
               #STATE_FAULT,
               #STATE_PROBLEM:
                   // The device is reachable, but faulty because of an error in a
                   // subordinated system --> check the modules
                   // Store the state of the different module in the diag DB
                   FOR #tempSlotIndex := 0 TO "USERDIAG_SLOTS_PER_DEVICE_UPPER_LIM" DO
                       IF (#ioSystemData.devices[#tempDeviceIndex].slots[#tempSlotIndex].configured = TRUE)
                       THEN
                           IF (#statDeviceProblemModules[#tempSlotIndex + 1] = TRUE)
                           THEN
                               // Problem in module
                               #ioSystemData.devices[#tempDeviceIndex].slots[#tempSlotIndex].faulty := FALSE;
                               #ioSystemData.devices[#tempDeviceIndex].slots[#tempSlotIndex].error := TRUE;
                               #ioSystemData.devices[#tempDeviceIndex].slots[#tempSlotIndex].problem := TRUE;
                               #ioSystemData.devices[#tempDeviceIndex].slots[#tempSlotIndex].state := #STATE_PROBLEM;

                               IF (#statDeviceFaultyModules[#tempSlotIndex + 1] = TRUE)
                               THEN
                                   // Fault in module
                                   #ioSystemData.devices[#tempDeviceIndex].slots[#tempSlotIndex].faulty := TRUE;
                                   #ioSystemData.devices[#tempDeviceIndex].slots[#tempSlotIndex].state := #STATE_FAULT;
                               END_IF;
                           ELSE
                               #ioSystemData.devices[#tempDeviceIndex].slots[#tempSlotIndex].error := FALSE;
                               #ioSystemData.devices[#tempDeviceIndex].slots[#tempSlotIndex].problem := FALSE;
                               #ioSystemData.devices[#tempDeviceIndex].slots[#tempSlotIndex].faulty := FALSE;
                           END_IF;

                           IF (#statDeviceExistingModules[#tempSlotIndex + 1] = TRUE)
                           THEN
                               // Module exists
                               #ioSystemData.devices[#tempDeviceIndex].slots[#tempSlotIndex].exists := TRUE;
                           ELSE
                               // Module does not exist
                               #ioSystemData.devices[#tempDeviceIndex].slots[#tempSlotIndex].exists := FALSE;
                           END_IF;
                       END_IF;
                   END_FOR;
               ELSE
                   // All modules are okay
                   FOR #tempSlotIndex := 0 TO "USERDIAG_SLOTS_PER_DEVICE_UPPER_LIM" DO
                       IF (#ioSystemData.devices[#tempDeviceIndex].slots[#tempSlotIndex].configured = TRUE)
                       THEN
                           #ioSystemData.devices[#tempDeviceIndex].slots[#tempSlotIndex].error := FALSE;
                           #ioSystemData.devices[#tempDeviceIndex].slots[#tempSlotIndex].problem := FALSE;
                           #ioSystemData.devices[#tempDeviceIndex].slots[#tempSlotIndex].faulty := FALSE;
                           #ioSystemData.devices[#tempDeviceIndex].slots[#tempSlotIndex].exists := TRUE;
                       END_IF;
                   END_FOR;
           END_CASE;
       END_IF;

       // Initialize the pointer for the next run
       #tempDeviceIndex := #ioSystemData.devices[#tempDeviceIndex].nextDevice;
   END_WHILE;


   // Write static values to outputs
   #error := #statError;
   #status := #statStatus;
   #statusID := #statStatusID;
END_FUNCTION_BLOCK

// folder: OBs

ORGANIZATION_BLOCK "Main"   // OB1, LAD, ProgramCycle
TITLE = "Main Program Sweep (Cycle)"
{ S7_Optimized_Access := 'TRUE' }
VERSION : 0.1
   VAR_INPUT
      Initial_Call : Bool;   // Initial call of this OB
      Remanence : Bool;   // =True, if remanent data are available
   END_VAR
BEGIN

REGION Network 1
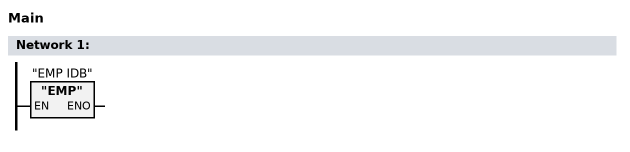
   RUNG wire#powerrail
      "EMP IDB"()
   END_RUNG
   // the same network as SCL:
   "EMP IDB"();   // "EMP"
END_REGION
END_ORGANIZATION_BLOCK

ORGANIZATION_BLOCK "Rack or station failure"   // OB86, LAD, RackStationFailure
{ S7_Optimized_Access := 'TRUE' }
VERSION : 0.1
   VAR_INPUT
      LADDR : Hw_Device;   // Hardware identifier
      Event_Class : Byte;   // Event class
      Fault_ID : Byte;   // Fault identifier
   END_VAR
BEGIN
END_ORGANIZATION_BLOCK

ORGANIZATION_BLOCK "Startup"   // OB100, LAD, Startup
TITLE = "Complete Restart"
{ S7_Optimized_Access := 'TRUE' }
VERSION : 0.1
// //============================================================================
// //SIEMENS AG
// //(c)Copyright 2017 All Rights Reserved
// //-----------------------------------------------------------------------------
// //Library: -
// //Tested with: S7-1516-3 PN/DP FW 2.5
// //Engineering: TIA Portal V15
// //Restrictions: -
// //Requirements: -
// //Functionality: Startup OB for Diagnostics
// //-----------------------------------------------------------------------------
// //Change log table:
// //Version  Date              Expert in charge                               Changes applied
// //01.00.00 25.04.2017 Siemens Industry Online Support First released version
// //============================================================================
   VAR_INPUT
      LostRetentive : Bool;   // True if retentive data are lost
      LostRTC : Bool;   // True if date and time are lost
   END_VAR
   VAR_TEMP
      index : Int;
   END_VAR
BEGIN

REGION Network 1: Set start user diagnostic
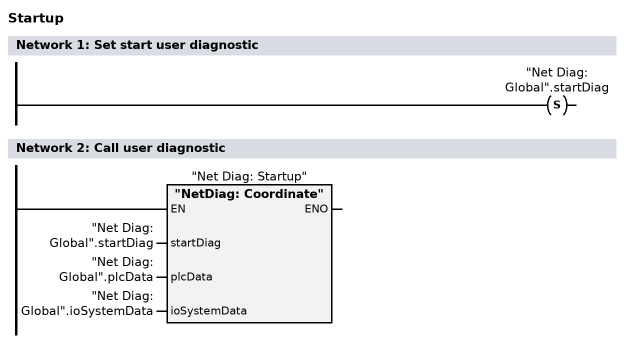
   RUNG wire#powerrail
      S_Coil( "Net Diag: Global".startDiag )
   END_RUNG
   // the same network as SCL:
   "Net Diag: Global".startDiag := TRUE;
END_REGION

REGION Network 2: Call user diagnostic
   RUNG wire#powerrail
      "Net Diag: Startup"(startDiag := "Net Diag: Global".startDiag, plcData := "Net Diag: Global".plcData, ioSystemData := "Net Diag: Global".ioSystemData)
   END_RUNG
   // the same network as SCL:
   "Net Diag: Startup"(startDiag := "Net Diag: Global".startDiag,   // "NetDiag: Coordinate"
                       plcData := "Net Diag: Global".plcData,
                       ioSystemData := "Net Diag: Global".ioSystemData);
END_REGION
END_ORGANIZATION_BLOCK

ORGANIZATION_BLOCK "Programming error"   // OB121, LAD, ProgrammingError
{ S7_Optimized_Access := 'TRUE' }
VERSION : 0.1
   VAR_INPUT
      BlockNr : UInt;   // Number of causing block
      Reaction : USInt;   // 0:ignore, 1:substitute, 2:skip
      Fault_ID : Byte;   // Fault identifier
      BlockType : USInt;   // 16#01:OB, 16#02:FC, 16#03:FB, 16#04:SFC, 16#05:SFB, 16#06:DB: Type of block causing the error
      Area : USInt;   // Area where the error occured
      DBNr : DB_ANY;   // DB number if Area = DB or DI
      Csg_OBNr : OB_Any;   // Number of OB causing the error
      Csg_Prio : USInt;   // Priority of OB causing the error
      Width : USInt;   // 0:bit, 1:byte, 2:word, 3:dword, 4:lword
   END_VAR
BEGIN
END_ORGANIZATION_BLOCK

ORGANIZATION_BLOCK "IO access error"   // OB122, LAD, IOAccessError
{ S7_Optimized_Access := 'TRUE' }
VERSION : 0.1
   VAR_INPUT
      BlockNr : UInt;   // Number of causing block
      Reaction : USInt;   // 0:ignore, 1:substitute, 2:skip
      Fault_ID : Byte;   // 16#42:reading, 16#43:writing
      BlockType : USInt;   // 16#01:OB, 16#02:FC, 16#03:FB, 16#04:SFC, 16#05:SFB, 16#06:DB: Type of block causing the error
      Area : USInt;   // 16#81:I, 16#82:Q: IO area where the IOaccess error occured
      DBNr : DB_ANY;   // Reserved for system
      Csg_OBNr : OB_Any;   // Number of OB causing the error
      Csg_Prio : USInt;   // Priority of OB causing the error
      Width : USInt;   // 0:bit, 1:byte, 2:word, 3:dword, 4:lword
   END_VAR
BEGIN
END_ORGANIZATION_BLOCK

// folder: Unsorted

FUNCTION_BLOCK "Code 128"   // FB2, SCL
{ S7_Optimized_Access := 'TRUE' }
VERSION : 0.1
   VAR_INPUT
      partNumber : String;
   END_VAR
   VAR_OUTPUT
      barcode : String;
   END_VAR
   VAR
      charsIn : Array[0..255] of Byte;
      charsOut : Array[0..255] of Byte;
      cnt : UInt;
      intVals : Array[0..255] of Int;
      sum : Int;
      checkSum : Int;
   END_VAR
   VAR_TEMP
      pn : String;
      i : Int;
   END_VAR
   VAR CONSTANT
      startChar : Char := 'Ì';
      stopChar : Char := 'Î';
   END_VAR
   // intVals[0] := 104;
BEGIN
   #pn := #partNumber;

   FOR #i := 0 TO 255 DO
       #charsIn[#i] := 16#00;
       #charsOut[#i] := 16#00;
       #intVals[#i] := 0;
   END_FOR;

   Strg_TO_Chars(Strg:=#pn,
                 pChars:=0,
                 Cnt=>#cnt,
                 Chars:=#charsIn);


   #sum := 104;
   FOR #i := 0 TO UINT_TO_INT(#cnt - 1) DO
       #intVals[#i] := CHAR_TO_INT(#charsIn[#i]) - 32;
       #intVals[#i] := #intVals[#i] * (#i + 1);
       #sum := #sum + #intVals[#i];
   END_FOR;
   #checkSum := (#sum MOD 103) + 32;
   IF #checkSum >= 127 THEN
       #checkSum := #checkSum + 68;
   END_IF;

   #charsOut[0] := #startChar;
   FOR #i := 1 TO UINT_TO_INT(#cnt) DO
       #charsOut[#i] := #charsIn[#i - 1];
   END_FOR;
   #charsOut[#cnt + 1] := INT_TO_BYTE(#checkSum);
   #charsOut[#cnt + 2] := INT_TO_BYTE(#stopChar);

   Chars_TO_Strg(Chars := #charsOut,
                 pChars := 0,
                 Cnt := #cnt + 3,
                 Strg => #barcode);
END_FUNCTION_BLOCK

FUNCTION_BLOCK "HMI Barcod Screen"   // FB3, SCL
{ S7_Optimized_Access := 'TRUE' }
VERSION : 0.1
   VAR_IN_OUT
      partCall : "Part Call Screen";
      barcodeScreen : "Barcode Screen";
      stations : "Stations";
   END_VAR
   VAR
      address : UInt;
      button : UInt;
      instCode128 : "Code 128";
      codeOut : String;
      pnOut : WString[40];
      station : UInt;
      oldSelectedRow : Int;
      oldOrderedBtn : Bool;
   END_VAR
   VAR_TEMP
      orderCancelled : Int;
      processedPN : String[40];
      selectedPN : String[40];
      userOrdered : Bool;
      selectedRow : Int;
      position : Int;
   END_VAR
   VAR CONSTANT
      maxRows : Int := 199;
   END_VAR
BEGIN
   REGION "GET USER ROW SELECTION"
       #selectedRow := "Get Part Call Row Number"(partCall := #partCall); 
   END_REGION

   REGION "ON SELECTION OF A PART CALL ROW
       IF #selectedRow <> 0 THEN
           IF #selectedRow <> #oldSelectedRow THEN

               REGION "GET BUTTON AND STATION NUMBERS"
                   #address := #partCall.row[#selectedRow - 1].address;
                   "Address to Station and Button"(address := #address,
                                                   station => #station,
                                                   button => #button);
               END_REGION

               REGION "CONVERT STRING TO BARCODE"

                   REGION "COPY TO LOCALS"
                       #selectedPN := WSTRING_TO_STRING(#partCall.row[#selectedRow - 1].tfPartNumber.value);
                   END_REGION

                   REGION "CHECK FOR MULTI LINE"

                       REGION "GET POSITON OF CARRIAGE RETURN"
                           #position := FIND(IN1 := #selectedPN, IN2 := '$L');
                       END_REGION

                       REGION "MULTILINE"
                           IF #position <> 0 THEN
                               #processedPN := LEFT(IN := #selectedPN, L := #position - 1);
                           END_IF;
                       END_REGION

                       REGION "SINGLE LINE"
                           IF #position = 0 THEN
                               #processedPN := #selectedPN;
                           END_IF;
                       END_REGION

                   END_REGION

                   REGION "CONVERT TO BARCODE"
                       #instCode128(partNumber := #processedPN,
                                    barcode => #codeOut);
                   END_REGION

                   REGION "OUTPUT FOR HMI SCREEN"
                       #barcodeScreen.partNumber := STRING_TO_WSTRING(#processedPN);
                       #barcodeScreen.barcode := #codeOut;
                   END_REGION

               END_REGION

           END_IF;
       END_IF;
   END_REGION

   REGION "PASS USER ORDERED"

       REGION "COPY TO LOCAL"
           #userOrdered := #barcodeScreen.ordered;
       END_REGION

       REGION "TURN OFF THE LIGHTS"
           #barcodeScreen.ordered := FALSE;
       END_REGION

       REGION "ON RISING EDGE"
           IF #userOrdered AND NOT #oldOrderedBtn THEN

               REGION "SET PART ORDERED"
                   #stations.me[#station - 1].partOrdered[#button - 1] := #userOrdered;
               END_REGION

           END_IF;
       END_REGION

       REGION "CHANGE DETECTION"
           #oldOrderedBtn := #userOrdered;
       END_REGION

   END_REGION

   REGION "CHANGE DETECTION"    
       #oldSelectedRow := #selectedRow;
   END_REGION
END_FUNCTION_BLOCK

FUNCTION_BLOCK "Initialize"   // FB4, SCL
{ S7_Optimized_Access := 'TRUE' }
VERSION : 0.1
   VAR_INPUT
      req : Bool;
   END_VAR
   VAR_IN_OUT
      stations : "Stations";
   END_VAR
   VAR
      rtElapsed : Real;
      rt : "Runtime Data";
   END_VAR
   VAR_TEMP
      i : Int;
      reset : Struct
         req : Bool;
         elapsed : Real;
      END_STRUCT;
      stnCount : Int;
      init : Bool;
   END_VAR
   VAR CONSTANT
      resetLimit : Real := 1.25;
   END_VAR
BEGIN
   REGION "GET STATION COUNT"
       #stnCount := "stnCount";
   END_REGION

   REGION "FIRST SCAN OR REQUEST"
       IF "FirstScan" OR #req THEN
           // initialize all stations on plc first scan
           FOR #i := 0 TO #stnCount DO
               #stations.me[#i].init.hard := TRUE;
           END_FOR;
       END_IF;
   END_REGION

   REGION "RUNTIME CALL"
       // get elapsed time
       #rt.elapsed := RUNTIME(#rt.mem);
       // convert to real data type
       #rtElapsed := LREAL_TO_REAL(#rt.elapsed);
   END_REGION

   REGION "BUTTON 0 BASED RESET TIMERS"
       FOR #i := 0 TO #stnCount DO

           REGION "PRE-CONDITION"
               // init off by default
               #init := FALSE;
               // request is button 0 on kp8
               #reset.req := #stations.me[#i].kp8In.%X0;
               // saved to shorter name
               #reset.elapsed := #stations.me[#i].elapsedTime.resetReq;
           END_REGION

           REGION "RESET REQUEST"
               IF NOT #reset.req THEN
                   #reset.elapsed := 0.0;
               END_IF;
               IF #reset.req THEN
                   // incriment elapsed time
                   #reset.elapsed := #reset.elapsed + #rtElapsed;
                   // timer expired condition
                   IF #reset.elapsed >= #resetLimit THEN
                       #init := TRUE;
                       #reset.elapsed := 0.0;
                   END_IF;
               END_IF;
               // save elapsed time
               #stations.me[#i].elapsedTime.resetReq := #reset.elapsed;
           END_REGION

           REGION "SAVE INITIALIZATIN REQUEST"
               #stations.me[#i].init.hard := #init;
           END_REGION

       END_FOR;
   END_REGION
END_FUNCTION_BLOCK

FUNCTION_BLOCK "Reset Init Requests"   // FB5, SCL
{ S7_Optimized_Access := 'TRUE' }
VERSION : 0.1
   VAR_IN_OUT
      stations : "Stations";
   END_VAR
   VAR
      placeHolder : Bool;
   END_VAR
   VAR_TEMP
      i : Int;
      stnCount : Int;
   END_VAR
BEGIN
   REGION "GET STATION COUNT"
       #stnCount := "stnCount";
   END_REGION

   REGION "RESET INITIALIZATION REQUESTS
       FOR #i := 0 TO #stnCount DO
           #stations.me[#i].init.hard := FALSE;
           #stations.me[#i].init.soft := FALSE;
       END_FOR;
   END_REGION
END_FUNCTION_BLOCK

FUNCTION_BLOCK "Record Part Request"   // FB6, SCL
{ S7_Optimized_Access := 'TRUE' }
VERSION : 0.1
   VAR_IN_OUT
      pRow : Int;
      requests : "Part Request Data";
      stations : "Stations";
   END_VAR
   VAR
      enterAddress : Bool;
      old : Struct
         presses : "Station Old Presses";
      END_STRUCT;
   END_VAR
   VAR_TEMP
      address : UInt;
      hasPart : Bool;
      i : Int;
      j : Int;
      k : Int;
      logAddress : UInt;
      noPart : Bool;
      oldPartReq : Bool;
      partReq : Bool;
      partNumber : WString;
      stnCount : Int;
      maxReqRows : Int;
   END_VAR
BEGIN
   REGION "COPY TO LOCAL"
       #maxReqRows := "partReqHmiRowCount";
       #stnCount := "stnCount";
   END_REGION

   REGION "FOR EACH STATION"
       FOR #i := 0 TO #stnCount DO

           REGION "FOR EACH BUTTON"
               // j = 0 is excluded because it is used as a station reset button
               FOR #j := 1 TO 7 DO

                   REGION "COPY TO LOCAL"
                       #partReq := #stations.me[#i].btnStates[#j];
                       #oldPartReq := #old.presses.me[#i,#j];
                   END_REGION

                   REGION "DETERMINE STATE"

                       REGION "ON NEW REQUEST"
                           IF #partReq AND NOT #oldPartReq THEN

                               REGION "SAVE FOR CHANGE DETECTION"
                                   #old.presses.me[#i, #j] := #stations.me[#i].btnStates[#j];
                               END_REGION

                               REGION "COPY TO LOCAL"
                                   #partNumber := #stations.me[#i].partNumbers[#j];
                               END_REGION

                               REGION "BUTTON HAS NO PN"
                                   IF LEN(#partNumber) = 0 THEN
                                       #hasPart := FALSE;
                                       #noPart := TRUE;
                                   END_IF;
                               END_REGION

                               REGION "BUTTON HAS PN"
                                   IF LEN(#partNumber) <> 0 THEN
                                       #hasPart := TRUE;
                                       #noPart := FALSE;
                                   END_IF;
                               END_REGION

                           END_IF;
                       END_REGION

                   END_REGION

                   REGION "NO PART"
                       IF #noPart THEN

                           REGION "TURN OFF THE LIGHTS"
                               #hasPart := FALSE;
                               #noPart := FALSE;
                               #enterAddress := FALSE;
                           END_REGION

                       END_IF;
                   END_REGION

                   REGION "HAS PART"
                       IF #hasPart THEN

                           REGION "TURN OFF THE LIGHTS"
                               #hasPart := FALSE;
                               #noPart := FALSE;
                               #enterAddress := FALSE;
                           END_REGION

                           REGION "CALCULATE ADDRESS"
                               #address := (INT_TO_UINT(#i) + 1) * 10 + (INT_TO_UINT(#j) + 1);
                           END_REGION

                           REGION "SET FLAG"
                               #enterAddress := TRUE;
                           END_REGION

                           REGION "CHECK FOR ENTRY IN DB"
                               REGION "FOR EACH ROW IN PART DB"
                                   FOR #k := 0 TO #maxReqRows DO

                                       REGION "COPY TO LOCAL"
                                           #logAddress := #requests.row[#k].address;
                                       END_REGION

                                       REGION "RESET FLAG"
                                           IF #logAddress = #address THEN
                                               #enterAddress := FALSE;
                                           END_IF;
                                       END_REGION

                                   END_FOR;
                               END_REGION
                           END_REGION


                       END_IF;
                   END_REGION

                   REGION "SAVE ROW DATA"
                       IF #enterAddress THEN

                           REGION "TURN OFF THE LIGHTS"
                               #enterAddress := FALSE;
                           END_REGION

                           REGION "ENTER PART REQUEST"
                               #stations.me[#i].partRequested[#j] := TRUE;
                           END_REGION

                           REGION "ADDRESS"
                               #requests.row[#pRow].address := #address;
                           END_REGION

                           REGION "LINE"
                               #requests.row[#pRow].tfLine.value := #stations.me[#i].line;
                           END_REGION

                           REGION "DROP ZONE"
                               #requests.row[#pRow].tfDropZone.value := USINT_TO_WSTRING(#stations.me[#i].dropZone);
                           END_REGION

                           REGION "PART NUMBER"
                               #requests.row[#pRow].tfPartNumber.value := #stations.me[#i].partNumbers[#j];
                           END_REGION

                           REGION "ELLAPSED TIME"
                               #requests.row[#pRow].tfTime.value := "Real to WString Timer"(#stations.me[#i].elapsedTime.partReq[#j]);
                           END_REGION

                           REGION "ROW POINTER"

                               REGION "INCREMENT"
                                   #pRow := #pRow + 1;
                               END_REGION

                               REGION "HIGH LIMIT ROLLOVER"
                                   IF #pRow > #maxReqRows THEN
                                       #pRow := 0;
                                   END_IF;
                               END_REGION

                           END_REGION

                       END_IF;
                   END_REGION

               END_FOR;
           END_REGION

       END_FOR;
   END_REGION
END_FUNCTION_BLOCK

FUNCTION_BLOCK "Part Timers"   // FB7, SCL
{ S7_Optimized_Access := 'TRUE' }
VERSION : 0.1
   VAR_IN_OUT
      stations : "Stations";
   END_VAR
   VAR
      rt : "Runtime Data";
      old : Struct
         presses : "Station Old Presses";
      END_STRUCT;
   END_VAR
   VAR_TEMP
      alottedTime : Real;
      btnCount : Int;
      elapsedTime : Real;
      i : Int;
      j : Int;
      partRequested : Bool;
      redTime : Real;
      remainingTime : Real;
      stnCount : Int;
      press : Struct
         current : Bool;
         old : Bool;
      END_STRUCT;
   END_VAR
BEGIN
   REGION "RUNTIME CALL"
       #rt.elapsed := RUNTIME(#rt.mem);
       #rt.asReal := LREAL_TO_REAL(#rt.elapsed);
   END_REGION

   REGION "COPY TO LOCAL"
       #stnCount := "stnCount";
       #btnCount := "ptsPerStn";
   END_REGION

   REGION "FOR EACH STATION"
       FOR #i := 0 TO #stnCount DO

           REGION "FOR EACH BUTTON"
               // j := 0 would be the reset button so it is skipped
               FOR #j := 1 TO #btnCount DO

                   REGION "RESET PART TIMER"

                       REGION "COPY TO LOCAL"
                           #press.current := #stations.me[#i].btnStates[#j];
                           #press.old := #old.presses.me[#i, #j];
                       END_REGION

                       REGION "ON PRESS FALLING EDGE"
                           IF NOT #press.current AND #press.old THEN
                               #stations.me[#i].elapsedTime.partReq[#j] := 0.0;
                           END_IF;
                           #old.presses.me[#i, #j] := #stations.me[#i].btnStates[#j];
                       END_REGION

                   END_REGION

                   REGION "PART REQUEST TIMER"

                       REGION "COPY TO LOCAL"
                           #partRequested := #stations.me[#i].btnStates[#j];
                       END_REGION

                       REGION "ON PART REQUEST"
                           IF #partRequested THEN

                               REGION "OUTPUT ELLAPSED TIME"
                                   // get saved time
                                   #elapsedTime := #stations.me[#i].elapsedTime.partReq[#j];
                                   // add elapsed time
                                   #elapsedTime += #rt.asReal;
                                   // save new value
                                   #stations.me[#i].elapsedTime.partReq[#j] := #elapsedTime;
                               END_REGION

                           END_IF;
                       END_REGION

                   END_REGION

               END_FOR;
           END_REGION

       END_FOR;
   END_REGION
END_FUNCTION_BLOCK

FUNCTION_BLOCK "Base Animations"   // FB8, SCL
{ S7_Optimized_Access := 'TRUE' }
VERSION : 0.1
   VAR_IN_OUT
      stations : "Stations";
   END_VAR
   VAR_TEMP
      animation : Int;
      i : Int;
      j : Int;
      partRequested : Bool;
      partOrdered : Bool;
      elapsedTime : Real;
      criticalTime : Real;
      alottedTime : Real;
      remainingTime : Real;
      stnCount : Int;
   END_VAR
   VAR CONSTANT
      anDefault : USInt := 0;
      anRequested : USInt := 1;
      anSolidRed : USInt := 2;
      anFlashRed : USInt := 3;
      anPartOrdered : USInt := 4;
   END_VAR
BEGIN
   REGION "COPY TO LOCAL"
       #stnCount := "stnCount";
   END_REGION

   REGION "FOR EACH STATION"
       FOR #i := 0 TO #stnCount DO

           REGION "FOR EACH BUTTON"
               // j := 0 would be the reset button so it is skipped
               FOR #j := 1 TO 7 DO

                   REGION "PART REQUEST TIMER"

                       REGION "COPY TO LOCAL"
                           #partRequested := #stations.me[#i].btnStates[#j];
                           #partOrdered := #stations.me[#i].partOrdered[#j];
                       END_REGION

                       REGION "PART REQUESTED"
                           IF #partRequested THEN

                               REGION "COPY TO LOCAL"
                                   // remaining time
                                   #elapsedTime := #stations.me[#i].elapsedTime.partReq[#j];
                                   #alottedTime := #stations.me[#i].presetTime.allotted[#j];
                                   #remainingTime := #alottedTime - #elapsedTime;
                                   // critical time
                                   #criticalTime := #stations.me[#i].presetTime.critical[#j];
                               END_REGION

                               REGION "DEFAULT ANIMATION STATE"
                                   IF #remainingTime > #criticalTime THEN
                                       #animation := #anRequested;
                                   END_IF;
                               END_REGION

                               REGION "ORDERED"
                                   IF #partOrdered THEN
                                       #animation := #anPartOrdered;
                                   END_IF;
                               END_REGION

                               REGION "SOLID RED ANIMATION STATE"
                                   IF #remainingTime <= #criticalTime AND #elapsedTime > 0.0 THEN
                                       #animation := #anSolidRed;
                                   END_IF;
                               END_REGION

                               REGION "FLASHING RED ANIMATION STATE
                                   IF #remainingTime <= 0.0 THEN
                                       #animation := #anFlashRed;
                                   END_IF;
                               END_REGION

                           END_IF;
                       END_REGION

                       REGION "PART NOT REQUESTED"
                           IF NOT #partRequested THEN
                               #animation := #anDefault;
                           END_IF;
                       END_REGION

                       REGION "OUTPUT"
                           #stations.me[#i].animations[#j] := #animation;
                       END_REGION

                   END_REGION

               END_FOR;
           END_REGION

       END_FOR;
   END_REGION
END_FUNCTION_BLOCK

FUNCTION_BLOCK "Format Part Call Requests"   // FB9, SCL
{ S7_Optimized_Access := 'TRUE' }
VERSION : 0.1
   VAR_IN_OUT
      requests : "Part Request Data";
      stations : "Stations";
   END_VAR
   VAR
      station : Int;
      button : Int;
   END_VAR
   VAR_TEMP
      address : Int;
      animate : USInt;
      maxRows : Int;
      timeAsReal : Real;
      timeAsTime : WString;
      i : Int;
      inStrRslt : Int;
      invisible : USInt;
      genericVisible : USInt;
      gray : USInt;
      darkGray : USInt;
      red : USInt;
      blue : USInt;
      redFlashing : USInt;
   END_VAR
   VAR CONSTANT
      visible : USInt := 1;
      anDefault : USInt := 0;
      anRequested : USInt := 1;
      anSolidRed : USInt := 2;
      anFlashRed : USInt := 3;
      anPartOrdered : USInt := 4;
   END_VAR
BEGIN
   REGION "COPY TO LOCAL"
       #invisible := "invisible";
       #maxRows := "partReqHmiRowCount";
       #gray := "BgGray";
       #darkGray := "disabled";
       #blue := "BgLBl";
       #red := "BgDRd";
       #redFlashing := "FlDrd";
   END_REGION


   REGION "ITERATE THROUGH VISIBLE TABLE ROWS"
       FOR #i := 0 TO #maxRows DO

           REGION "COPY TO LOCAL"
               #address := UINT_TO_INT(#requests.row[#i].address);
           END_REGION

           REGION "HIDE UNPOPULATED ROWS"
               IF #address = 0 THEN
                   #requests.row[#i].pbSelection.animate := #invisible;
                   #requests.row[#i].rtBackground.animate := #invisible;
                   #animate := 0;
                   #requests.row[#i].tfDropZone.animate := #invisible;
                   #requests.row[#i].tfLine.animate := #invisible;
                   #requests.row[#i].tfPartNumber.animateSL := #invisible;
                   #requests.row[#i].tfPartNumber.animateDL := #invisible;
                   #requests.row[#i].tfTime.animate := #invisible;
               END_IF;
           END_REGION

           REGION "ANIMATE POPULATED ROWS"

               REGION "ANIMATE ROWS WITH DATA"
                   IF #address <> 0 THEN

                       REGION "GET POINTERS FOR STATION ARRAY"
                           #station := #address / 10 - 1;
                           #button := #address MOD 10 - 1;
                       END_REGION

                       REGION "SET ANIMATE"
                           CASE #stations.me[#station].animations[#button] OF
                               #anRequested:
                                   #animate := #gray;
                               #anSolidRed:
                                   #animate := #red;
                               #anFlashRed:
                                   #animate := #redFlashing;
                               #anPartOrdered:
                                   #animate := #blue;
                               ELSE
                                   #animate := #invisible;
                           END_CASE;
                       END_REGION


                       REGION "ANIMATIONS"

                           REGION "PUSHBUTTON VISIBILITY"
                               #requests.row[#i].pbSelection.animate := #visible;
                           END_REGION

                           REGION "BACKGROUND VISIBILITY"
                               #requests.row[#i].rtBackground.animate := #darkGray;
                           END_REGION

                           REGION "DROP ZONE" 
                               #requests.row[#i].tfDropZone.animate := #animate;
                               #requests.row[#i].tfDropZone.value := "Strip Sign"(UINT_TO_WSTRING(#stations.me[#station].dropZone));
                           END_REGION

                           REGION "LINE"
                               #requests.row[#i].tfLine.animate := #animate;
                               #requests.row[#i].tfLine.value := #stations.me[#station].line;
                           END_REGION

                           REGION "PART NUMBER"
                               #requests.row[#i].tfPartNumber.animateSL := #animate;
                               #requests.row[#i].tfPartNumber.value := #stations.me[#station].partNumbers[#button];
                               REGION "DETERMINE VISIBLE ROWS"

                                   REGION "FIND CARRIAGE RETURN"
                                       #inStrRslt := FIND(IN1 := #requests.row[#i].tfPartNumber.value,
                                                          IN2 := wstring#'$L');
                                   END_REGION

                                   REGION "SINGLE LINE"
                                       IF #inStrRslt = 0 THEN
                                           #requests.row[#i].tfPartNumber.animateSL := #animate;
                                           #requests.row[#i].tfPartNumber.animateDL := #invisible;
                                       END_IF;
                                   END_REGION

                                   REGION "DOUBLE LINE"
                                       IF #inStrRslt <> 0 THEN
                                           #requests.row[#i].tfPartNumber.animateSL := #invisible;
                                           #requests.row[#i].tfPartNumber.animateDL := #animate;
                                       END_IF;
                                   END_REGION

                               END_REGION

                           END_REGION

                           REGION "TIME"
                               #requests.row[#i].tfTime.animate := #animate;
                               #timeAsReal := #stations.me[#station].presetTime.allotted[#button];
                               #timeAsReal -= #stations.me[#station].elapsedTime.partReq[#button];
                               #requests.row[#i].tfTime.value := "Real to WString Timer"(#timeAsReal);
                           END_REGION

                       END_REGION

                   END_IF;
               END_REGION

           END_REGION

       END_FOR;
   END_REGION
END_FUNCTION_BLOCK

FUNCTION_BLOCK "KP8 Expanded Animations"   // FB10, SCL
{ S7_Optimized_Access := 'TRUE' }
VERSION : 0.1
   VAR_IN_OUT
      stations : "Stations";
   END_VAR
   VAR_TEMP
      i : Int;
      j : Int;
      colorBox : DWord;
      animation : Int;
      mask : DWord;
   END_VAR
   VAR CONSTANT
      stationCount : Int := 23;
      buttonCount : Int := 7;
      anSolidRed : USInt := 2;
      anFlashRed : USInt := 3;
      anBlue : USInt := 4;
   END_VAR
BEGIN
   REGION "LOOP THROUGH STATIONS"
       FOR #i := 0 TO #stationCount DO

           REGION "LOOP THROUGH BUTTONS"
               FOR #j := 0 TO #buttonCount DO

                   REGION "GET ANIMATION"
                       #animation := #stations.me[#i].animations[#j];
                   END_REGION

                   REGION "SOLID RED"
                       IF #animation = #anSolidRed THEN
                           #colorBox := #stations.me[#i].kp8Out;
                           #mask := 16#FEFEFEFF;
                           #mask := ROL_DWORD(IN := #mask,
                                                 N := INT_TO_UINT(#j));
                           #colorBox := #colorBox AND #mask;
                           #mask := 16#100_0000;
                           #mask := ROL_DWORD(IN := #mask,
                                                 N := INT_TO_UINT(#j));
                           #colorBox := #colorBox OR #mask;
                           #stations.me[#i].kp8Out := #colorBox;
                       END_IF;
                   END_REGION

                   REGION "FLASHING RED"
                       IF #animation = #anFlashRed THEN

                           REGION "RED ON"
                               IF "Clock_1Hz" THEN
                                   #colorBox := #stations.me[#i].kp8Out;
                                   #mask := 16#FEFEFEFF;
                                   #mask := ROL_DWORD(IN := #mask,
                                                         N := INT_TO_UINT(#j));
                                   #colorBox := #colorBox AND #mask;
                                   #mask := 16#100_0000;
                                   #mask := ROL_DWORD(IN := #mask,
                                                         N := INT_TO_UINT(#j));
                                   #colorBox := #colorBox OR #mask;
                                   #stations.me[#i].kp8Out := #colorBox;
                               END_IF;
                           END_REGION

                           REGION "RED OFF"
                               IF NOT "Clock_1Hz" THEN
                                   #colorBox := #stations.me[#i].kp8Out;
                                   #mask := 16#FEFEFEFF;
                                   #mask := ROL_DWORD(IN := #mask,
                                                         N := INT_TO_UINT(#j));
                                   #colorBox := #colorBox AND #mask;
                                   #stations.me[#i].kp8Out := #colorBox;
                               END_IF;
                           END_REGION

                       END_IF;
                   END_REGION

                   REGION "BLUE"
                       IF #animation = #anBlue THEN
                           #colorBox := #stations.me[#i].kp8Out;
                           #mask := 16#FEFEFEFF;
                           #mask := ROL_DWORD(IN := #mask,
                                              N := INT_TO_UINT(#j));
                           #colorBox := #colorBox AND #mask;
                           #mask := 16#0000_0100;
                           #mask := ROL_DWORD(IN := #mask,
                                                 N := INT_TO_UINT(#j));
                           #colorBox := #colorBox OR #mask;
                           #stations.me[#i].kp8Out := #colorBox;
                       END_IF;
                   END_REGION

               END_FOR;
           END_REGION

       END_FOR;
   END_REGION
END_FUNCTION_BLOCK

FUNCTION_BLOCK "Stack Light Animations"   // FB11, SCL
{ S7_Optimized_Access := 'TRUE' }
VERSION : 0.1
   VAR_IN_OUT
      stations : "Stations";
   END_VAR
   VAR_TEMP
      animation : Int;
      i : Int;
      j : Int;
      stackLight : DWord;
   END_VAR
   VAR CONSTANT
      anDefault : USInt := 0;
      anRequested : USInt := 1;
      anSolidRed : USInt := 2;
      anFlashRed : USInt := 3;
      anPartOrdered : USInt := 4;
      buttonCount : Int := 7;
      "Part 01" : Int := 7;
      "Part 01 Green On" : DWord := 16#0400_0000;
      "Part 01 Red On" : DWord := 16#0100_0000;
      "Part 01 Yellow On" : DWord := 16#0200_0000;
      "Part 02" : Int := 3;
      "Part 02 Green On" : DWord := 16#2000_0000;
      "Part 02 Red On" : DWord := 16#0800_0000;
      "Part 02 Yellow On" : DWord := 16#1000_0000;
      "Part 03" : Int := 6;
      "Part 03 Green On" : DWord := 16#0001_0000;
      "Part 03 Red On" : DWord := 16#4000_0000;
      "Part 03 Yellow On" : DWord := 16#8000_0000;
      "Part 04" : Int := 2;
      "Part 04 Green On" : DWord := 16#0008_0000;
      "Part 04 Yellow On" : DWord := 16#0004_0000;
      "Part 04 Red On" : DWord := 16#0002_0000;
      "Part 05" : Int := 5;
      "Part 05 Green On" : DWord := 16#0040_0000;
      "Part 05 Red On" : DWord := 16#0010_0000;
      "Part 05 Yellow On" : DWord := 16#0020_0000;
      "Part 06" : Int := 1;
      "Part 06 Green On" : DWord := 16#0000_0200;
      "Part 06 Red On" : DWord := 16#0080_0000;
      "Part 06 Yellow On" : DWord := 16#0000_0100;
      stationCount : Int := 23;
   END_VAR
BEGIN
   REGION "LOOP THROUGH STATIONS"
       FOR #i := 0 TO #stationCount DO

           REGION "LOOP THROUGH BUTTONS"
               FOR #j := 0 TO #buttonCount DO

                   REGION "COPY INTO LOCAL"
                       #stackLight := #stations.me[#i].stackLightOut;
                       #animation := #stations.me[#i].animations[#j];
                   END_REGION

                   REGION "GREEN"
                       IF #animation = #anDefault THEN
                           CASE #j OF
                               #"Part 01":
                                   #stackLight := #stackLight AND (NOT #"Part 01 Red On");
                                   #stackLight := #stackLight AND (NOT #"Part 01 Yellow On");
                                   #stackLight := #stackLight OR #"Part 01 Green On";
                               #"Part 02":
                                   #stackLight := #stackLight AND (NOT #"Part 02 Red On");
                                   #stackLight := #stackLight AND (NOT #"Part 02 Yellow On");
                                   #stackLight := #stackLight OR #"Part 02 Green On";
                               #"Part 03":
                                   #stackLight := #stackLight AND (NOT #"Part 03 Red On");
                                   #stackLight := #stackLight AND (NOT #"Part 03 Yellow On");
                                   #stackLight := #stackLight OR #"Part 03 Green On";
                               #"Part 04":
                                   #stackLight := #stackLight AND (NOT #"Part 04 Red On");
                                   #stackLight := #stackLight AND (NOT #"Part 04 Yellow On");
                                   #stackLight := #stackLight OR #"Part 04 Green On";
                               #"Part 05":
                                   #stackLight := #stackLight AND (NOT #"Part 05 Red On");
                                   #stackLight := #stackLight AND (NOT #"Part 05 Yellow On");
                                   #stackLight := #stackLight OR #"Part 05 Green On";
                               #"Part 06":
                                   #stackLight := #stackLight AND (NOT #"Part 06 Red On");
                                   #stackLight := #stackLight AND (NOT #"Part 06 Yellow On");
                                   #stackLight := #stackLight OR #"Part 06 Green On";
                               ELSE
                                   ;
                           END_CASE;
                       END_IF;
                   END_REGION

                   REGION "YELLOW"
                       IF #animation = #anRequested THEN
                           CASE #j OF
                               #"Part 01":
                                   #stackLight := #stackLight AND (NOT #"Part 01 Red On");
                                   #stackLight := #stackLight OR #"Part 01 Yellow On";
                                   #stackLight := #stackLight AND (NOT #"Part 01 Green On");
                               #"Part 02":
                                   #stackLight := #stackLight AND (NOT #"Part 02 Red On");
                                   #stackLight := #stackLight OR #"Part 02 Yellow On";
                                   #stackLight := #stackLight AND (NOT #"Part 02 Green On");
                               #"Part 03":
                                   #stackLight := #stackLight AND (NOT #"Part 03 Red On");
                                   #stackLight := #stackLight OR #"Part 03 Yellow On";
                                   #stackLight := #stackLight AND (NOT #"Part 03 Green On");
                               #"Part 04":
                                   #stackLight := #stackLight AND (NOT #"Part 04 Red On");
                                   #stackLight := #stackLight OR #"Part 04 Yellow On";
                                   #stackLight := #stackLight AND (NOT #"Part 04 Green On");
                               #"Part 05":
                                   #stackLight := #stackLight AND (NOT #"Part 05 Red On");
                                   #stackLight := #stackLight OR #"Part 05 Yellow On";
                                   #stackLight := #stackLight AND (NOT #"Part 05 Green On");
                               #"Part 06":
                                   #stackLight := #stackLight AND (NOT #"Part 06 Red On");
                                   #stackLight := #stackLight OR #"Part 06 Yellow On";
                                   #stackLight := #stackLight AND (NOT #"Part 06 Green On");
                               ELSE
                                   ;
                           END_CASE;
                       END_IF;
                   END_REGION

                   REGION "SOLID RED"
                       IF #animation = #anSolidRed THEN
                           CASE #j OF
                               #"Part 01":
                                   #stackLight := #stackLight OR #"Part 01 Red On";
                                   #stackLight := #stackLight AND (NOT #"Part 01 Yellow On");
                                   #stackLight := #stackLight AND (NOT #"Part 01 Green On");
                               #"Part 02":
                                   #stackLight := #stackLight OR #"Part 02 Red On";
                                   #stackLight := #stackLight AND (NOT #"Part 02 Yellow On");
                                   #stackLight := #stackLight AND (NOT #"Part 02 Green On");
                               #"Part 03":
                                   #stackLight := #stackLight OR #"Part 03 Red On";
                                   #stackLight := #stackLight AND (NOT #"Part 03 Yellow On");
                                   #stackLight := #stackLight AND (NOT #"Part 03 Green On");
                               #"Part 04":
                                   #stackLight := #stackLight OR #"Part 04 Red On";
                                   #stackLight := #stackLight AND (NOT #"Part 04 Yellow On");
                                   #stackLight := #stackLight AND (NOT #"Part 04 Green On");
                               #"Part 05":
                                   #stackLight := #stackLight OR #"Part 05 Red On";
                                   #stackLight := #stackLight AND (NOT #"Part 05 Yellow On");
                                   #stackLight := #stackLight AND (NOT #"Part 05 Green On");
                               #"Part 06":
                                   #stackLight := #stackLight OR #"Part 06 Red On";
                                   #stackLight := #stackLight AND (NOT #"Part 06 Yellow On");
                                   #stackLight := #stackLight AND (NOT #"Part 06 Green On");
                               ELSE
                                   ;
                           END_CASE;
                       END_IF;
                   END_REGION

                   REGION "FLASHING RED"
                       IF #animation = #anFlashRed THEN

                           REGION "RED ON"
                               IF "Clock_1Hz" THEN
                                   CASE #j OF
                                       #"Part 01":
                                           #stackLight := #stackLight OR #"Part 01 Red On";
                                           #stackLight := #stackLight AND (NOT #"Part 01 Yellow On");
                                           #stackLight := #stackLight AND (NOT #"Part 01 Green On");
                                       #"Part 02":
                                           #stackLight := #stackLight OR #"Part 02 Red On";
                                           #stackLight := #stackLight AND (NOT #"Part 02 Yellow On");
                                           #stackLight := #stackLight AND (NOT #"Part 02 Green On");
                                       #"Part 03":
                                           #stackLight := #stackLight OR #"Part 03 Red On";
                                           #stackLight := #stackLight AND (NOT #"Part 03 Yellow On");
                                           #stackLight := #stackLight AND (NOT #"Part 03 Green On");
                                       #"Part 04":
                                           #stackLight := #stackLight OR #"Part 04 Red On";
                                           #stackLight := #stackLight AND (NOT #"Part 04 Yellow On");
                                           #stackLight := #stackLight AND (NOT #"Part 04 Green On");
                                       #"Part 05":
                                           #stackLight := #stackLight OR #"Part 05 Red On";
                                           #stackLight := #stackLight AND (NOT #"Part 05 Yellow On");
                                           #stackLight := #stackLight AND (NOT #"Part 05 Green On");
                                       #"Part 06":
                                           #stackLight := #stackLight OR #"Part 06 Red On";
                                           #stackLight := #stackLight AND (NOT #"Part 06 Yellow On");
                                           #stackLight := #stackLight AND (NOT #"Part 06 Green On");
                                       ELSE
                                           ;
                                   END_CASE;
                               END_IF;
                           END_REGION

